REGION Network 75
   RUNG wire#powerrail
      Contact( "LimiteMantBoost2" )
      Coil( "DB32".Static_194 )
   END_RUNG
   // the same network as SCL:
   "DB32".Static_194 := "LimiteMantBoost2";
END_REGION

REGION Network 76
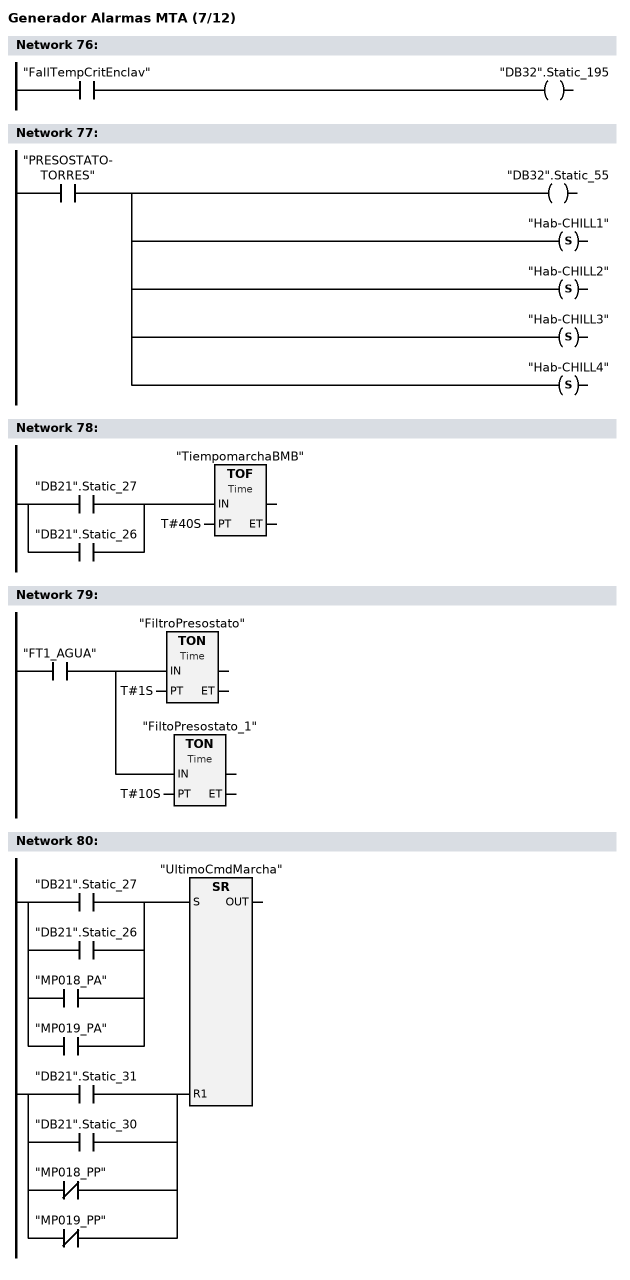
   RUNG wire#powerrail
      Contact( "FallTempCritEnclav" )
      Coil( "DB32".Static_195 )
   END_RUNG
   // the same network as SCL:
   "DB32".Static_195 := "FallTempCritEnclav";
END_REGION

REGION Network 77
   RUNG wire#powerrail
      Contact( "PRESOSTATO-TORRES" )
      wire#w1
      Coil( "DB32".Static_55 )
   END_RUNG
   RUNG wire#w1
      S_Coil( "Hab-CHILL1" )
   END_RUNG
   RUNG wire#w1
      S_Coil( "Hab-CHILL2" )
   END_RUNG
   RUNG wire#w1
      S_Coil( "Hab-CHILL3" )
   END_RUNG
   RUNG wire#w1
      S_Coil( "Hab-CHILL4" )
   END_RUNG
   // the same network as SCL:
   "DB32".Static_55 := "PRESOSTATO-TORRES";
   IF "PRESOSTATO-TORRES" THEN
       "Hab-CHILL1" := TRUE;
       "Hab-CHILL2" := TRUE;
       "Hab-CHILL3" := TRUE;
       "Hab-CHILL4" := TRUE;
   END_IF;
END_REGION

REGION Network 78
   "TiempomarchaBMB".TOF(in := "DB21".Static_27 OR "DB21".Static_26, pt := T#40S);
END_REGION

REGION Network 79
   "FiltroPresostato".TON(pt := T#1S, in := "FT1_AGUA");
   "FiltoPresostato_1".TON(pt := T#10S, in := "FT1_AGUA");
END_REGION

REGION Network 80
   RUNG wire#powerrail
      Contact( "DB21".Static_27 )
      wire#w1
      S_SR(operand := "UltimoCmdMarcha", r1 := wire#w2)
   END_RUNG
   RUNG wire#powerrail
      Contact( "DB21".Static_26 )
   END_RUNG wire#w1
   RUNG wire#powerrail
      Contact( "MP018_PA" )
   END_RUNG wire#w1
   RUNG wire#powerrail
      Contact( "MP019_PA" )
   END_RUNG wire#w1
   RUNG wire#powerrail
      Contact( "DB21".Static_31 )
   END_RUNG wire#w2
   RUNG wire#powerrail
      Contact( "DB21".Static_30 )
   END_RUNG wire#w2
   RUNG wire#powerrail
      I_Contact( "MP018_PP" )
   END_RUNG wire#w2
   RUNG wire#powerrail
      I_Contact( "MP019_PP" )
   END_RUNG wire#w2
   // the same network as SCL:
   IF "DB21".Static_27 OR "DB21".Static_26 OR "MP018_PA" OR "MP019_PA" THEN
       "UltimoCmdMarcha" := TRUE;   // SR flip-flop
   END_IF;
   IF "DB21".Static_31 OR "DB21".Static_30 OR NOT "MP018_PP" OR NOT "MP019_PP" THEN
       "UltimoCmdMarcha" := FALSE;
   END_IF;
END_REGION

REGION Network 81
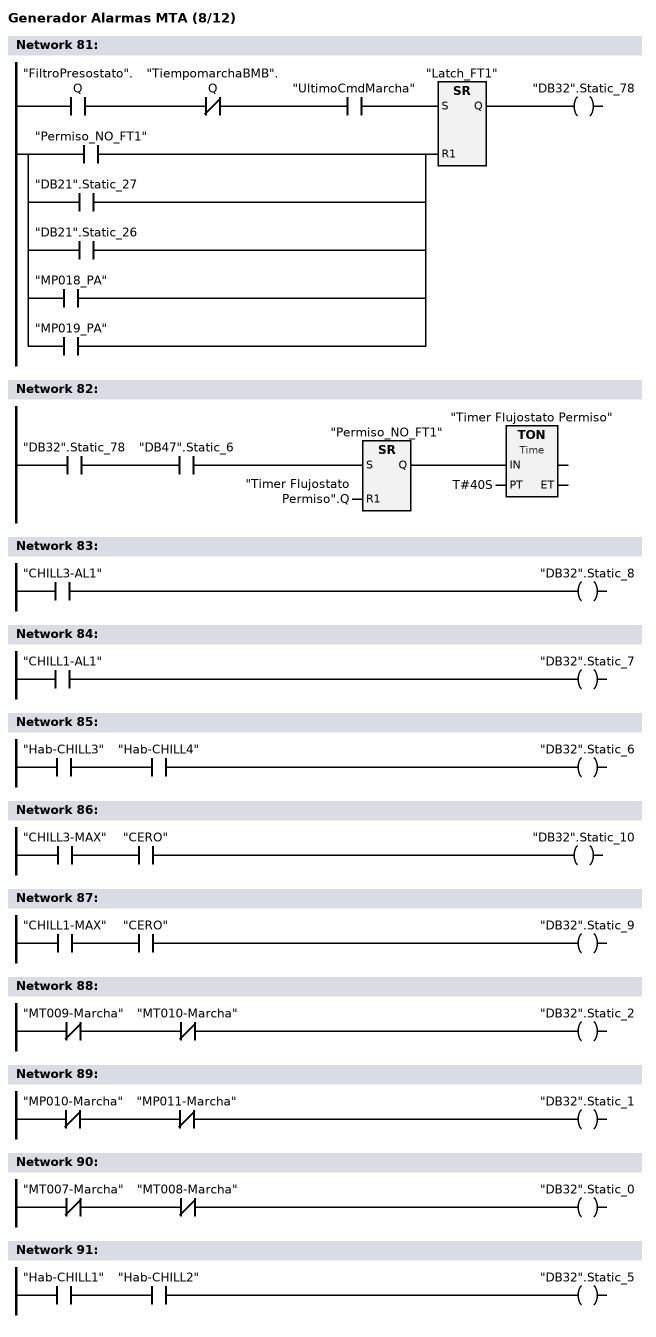
   RUNG wire#powerrail
      Contact( "FiltroPresostato".Q )
      I_Contact( "TiempomarchaBMB".Q )
      Contact( "UltimoCmdMarcha" )
      S_SR(operand := "Latch_FT1", r1 := wire#w1)
      Coil( "DB32".Static_78 )
   END_RUNG
   RUNG wire#powerrail
      Contact( "Permiso_NO_FT1" )
   END_RUNG wire#w1
   RUNG wire#powerrail
      Contact( "DB21".Static_27 )
   END_RUNG wire#w1
   RUNG wire#powerrail
      Contact( "DB21".Static_26 )
   END_RUNG wire#w1
   RUNG wire#powerrail
      Contact( "MP018_PA" )
   END_RUNG wire#w1
   RUNG wire#powerrail
      Contact( "MP019_PA" )
   END_RUNG wire#w1
   // the same network as SCL:
   IF "FiltroPresostato".Q AND NOT "TiempomarchaBMB".Q AND "UltimoCmdMarcha" THEN
       "Latch_FT1" := TRUE;   // SR flip-flop
   END_IF;
   IF "Permiso_NO_FT1" OR "DB21".Static_27 OR "DB21".Static_26 OR "MP018_PA" OR "MP019_PA" THEN
       "Latch_FT1" := FALSE;
   END_IF;
   "DB32".Static_78 := "Latch_FT1";
END_REGION

REGION Network 82
   IF "DB32".Static_78 AND "DB47".Static_6 THEN
       "Permiso_NO_FT1" := TRUE;   // SR flip-flop
   END_IF;
   IF "Timer Flujostato Permiso".Q THEN "Permiso_NO_FT1" := FALSE; END_IF;
   "Timer Flujostato Permiso".TON(in := "Permiso_NO_FT1", pt := T#40S);
END_REGION

REGION Network 83
   RUNG wire#powerrail
      Contact( "CHILL3-AL1" )
      Coil( "DB32".Static_8 )
   END_RUNG
   // the same network as SCL:
   "DB32".Static_8 := "CHILL3-AL1";
END_REGION

REGION Network 84
   RUNG wire#powerrail
      Contact( "CHILL1-AL1" )
      Coil( "DB32".Static_7 )
   END_RUNG
   // the same network as SCL:
   "DB32".Static_7 := "CHILL1-AL1";
END_REGION

REGION Network 85
   RUNG wire#powerrail
      Contact( "Hab-CHILL3" )
      Contact( "Hab-CHILL4" )
      Coil( "DB32".Static_6 )
   END_RUNG
   // the same network as SCL:
   "DB32".Static_6 := "Hab-CHILL3" AND "Hab-CHILL4";
END_REGION

REGION Network 86
   RUNG wire#powerrail
      Contact( "CHILL3-MAX" )
      Contact( "CERO" )
      Coil( "DB32".Static_10 )
   END_RUNG
   // the same network as SCL:
   "DB32".Static_10 := "CHILL3-MAX" AND "CERO";
END_REGION

REGION Network 87
   RUNG wire#powerrail
      Contact( "CHILL1-MAX" )
      Contact( "CERO" )
      Coil( "DB32".Static_9 )
   END_RUNG
   // the same network as SCL:
   "DB32".Static_9 := "CHILL1-MAX" AND "CERO";
END_REGION

REGION Network 88
   RUNG wire#powerrail
      I_Contact( "MT009-Marcha" )
      I_Contact( "MT010-Marcha" )
      Coil( "DB32".Static_2 )
   END_RUNG
   // the same network as SCL:
   "DB32".Static_2 := NOT "MT009-Marcha" AND NOT "MT010-Marcha";
END_REGION

REGION Network 89
   RUNG wire#powerrail
      I_Contact( "MP010-Marcha" )
      I_Contact( "MP011-Marcha" )
      Coil( "DB32".Static_1 )
   END_RUNG
   // the same network as SCL:
   "DB32".Static_1 := NOT "MP010-Marcha" AND NOT "MP011-Marcha";
END_REGION

REGION Network 90
   RUNG wire#powerrail
      I_Contact( "MT007-Marcha" )
      I_Contact( "MT008-Marcha" )
      Coil( "DB32".Static_0 )
   END_RUNG
   // the same network as SCL:
   "DB32".Static_0 := NOT "MT007-Marcha" AND NOT "MT008-Marcha";
END_REGION

REGION Network 91
   RUNG wire#powerrail
      Contact( "Hab-CHILL1" )
      Contact( "Hab-CHILL2" )
      Coil( "DB32".Static_5 )
   END_RUNG
   // the same network as SCL:
   "DB32".Static_5 := "Hab-CHILL1" AND "Hab-CHILL2";
END_REGION

REGION Network 92
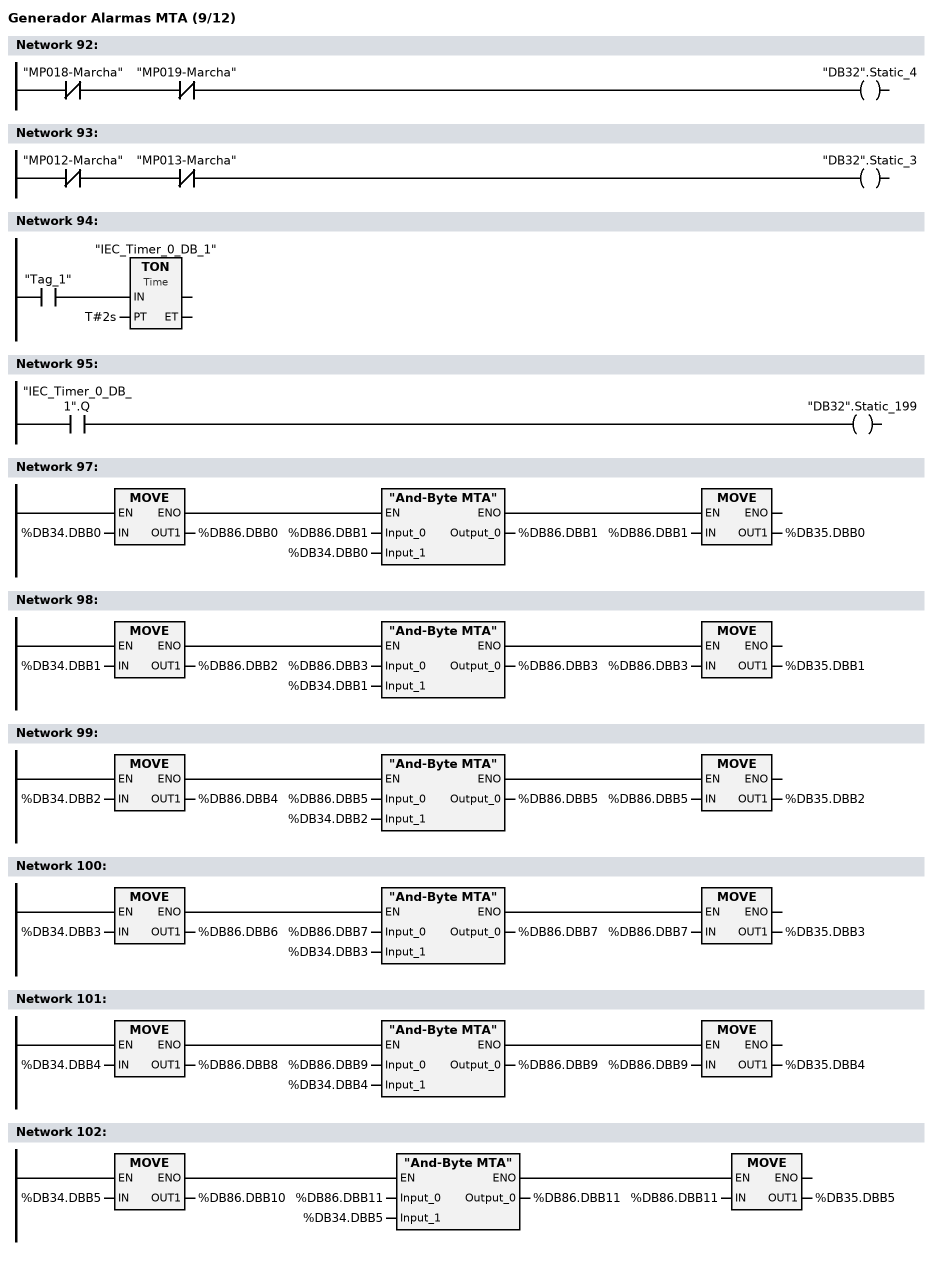
   RUNG wire#powerrail
      I_Contact( "MP018-Marcha" )
      I_Contact( "MP019-Marcha" )
      Coil( "DB32".Static_4 )
   END_RUNG
   // the same network as SCL:
   "DB32".Static_4 := NOT "MP018-Marcha" AND NOT "MP019-Marcha";
END_REGION

REGION Network 93
   RUNG wire#powerrail
      I_Contact( "MP012-Marcha" )
      I_Contact( "MP013-Marcha" )
      Coil( "DB32".Static_3 )
   END_RUNG
   // the same network as SCL:
   "DB32".Static_3 := NOT "MP012-Marcha" AND NOT "MP013-Marcha";
END_REGION

REGION Network 94
   "IEC_Timer_0_DB_1".TON(IN := "Tag_1", PT := T#2s);
END_REGION

REGION Network 95
   RUNG wire#powerrail
      Contact( "IEC_Timer_0_DB_1".Q )
      Coil( "DB32".Static_199 )
   END_RUNG
   // the same network as SCL:
   "DB32".Static_199 := "IEC_Timer_0_DB_1".Q;
END_REGION

REGION Network 97
   RUNG wire#powerrail
      { S7_GenerateENO := "TRUE" } Move(in := %DB34.DBB0, out1 => %DB86.DBB0)
      "And-Byte MTA"(Input_0 := %DB86.DBB1, Input_1 := %DB34.DBB0, Output_0 => %DB86.DBB1)
      { S7_GenerateENO := "TRUE" } Move(in := %DB86.DBB1, out1 => %DB35.DBB0)
   END_RUNG
   // the same network as SCL:
   // ENO of a box is taken as its EN; it also drops when the box reports an error
   %DB86.DBB0 := %DB34.DBB0;
   "And-Byte MTA"(Input_0 := %DB86.DBB1, Input_1 := %DB34.DBB0, Output_0 => %DB86.DBB1, ENO => #_w1);
   IF #_w1 THEN %DB35.DBB0 := %DB86.DBB1; END_IF;
END_REGION

REGION Network 98
   RUNG wire#powerrail
      { S7_GenerateENO := "TRUE" } Move(in := %DB34.DBB1, out1 => %DB86.DBB2)
      "And-Byte MTA"(Input_0 := %DB86.DBB3, Input_1 := %DB34.DBB1, Output_0 => %DB86.DBB3)
      { S7_GenerateENO := "TRUE" } Move(in := %DB86.DBB3, out1 => %DB35.DBB1)
   END_RUNG
   // the same network as SCL:
   // ENO of a box is taken as its EN; it also drops when the box reports an error
   %DB86.DBB2 := %DB34.DBB1;
   "And-Byte MTA"(Input_0 := %DB86.DBB3, Input_1 := %DB34.DBB1, Output_0 => %DB86.DBB3, ENO => #_w1);
   IF #_w1 THEN %DB35.DBB1 := %DB86.DBB3; END_IF;
END_REGION

REGION Network 99
   RUNG wire#powerrail
      { S7_GenerateENO := "TRUE" } Move(in := %DB34.DBB2, out1 => %DB86.DBB4)
      "And-Byte MTA"(Input_0 := %DB86.DBB5, Input_1 := %DB34.DBB2, Output_0 => %DB86.DBB5)
      { S7_GenerateENO := "TRUE" } Move(in := %DB86.DBB5, out1 => %DB35.DBB2)
   END_RUNG
   // the same network as SCL:
   // ENO of a box is taken as its EN; it also drops when the box reports an error
   %DB86.DBB4 := %DB34.DBB2;
   "And-Byte MTA"(Input_0 := %DB86.DBB5, Input_1 := %DB34.DBB2, Output_0 => %DB86.DBB5, ENO => #_w1);
   IF #_w1 THEN %DB35.DBB2 := %DB86.DBB5; END_IF;
END_REGION

REGION Network 100
   RUNG wire#powerrail
      { S7_GenerateENO := "TRUE" } Move(in := %DB34.DBB3, out1 => %DB86.DBB6)
      "And-Byte MTA"(Input_0 := %DB86.DBB7, Input_1 := %DB34.DBB3, Output_0 => %DB86.DBB7)
      { S7_GenerateENO := "TRUE" } Move(in := %DB86.DBB7, out1 => %DB35.DBB3)
   END_RUNG
   // the same network as SCL:
   // ENO of a box is taken as its EN; it also drops when the box reports an error
   %DB86.DBB6 := %DB34.DBB3;
   "And-Byte MTA"(Input_0 := %DB86.DBB7, Input_1 := %DB34.DBB3, Output_0 => %DB86.DBB7, ENO => #_w1);
   IF #_w1 THEN %DB35.DBB3 := %DB86.DBB7; END_IF;
END_REGION

REGION Network 101
   RUNG wire#powerrail
      { S7_GenerateENO := "TRUE" } Move(in := %DB34.DBB4, out1 => %DB86.DBB8)
      "And-Byte MTA"(Input_0 := %DB86.DBB9, Input_1 := %DB34.DBB4, Output_0 => %DB86.DBB9)
      { S7_GenerateENO := "TRUE" } Move(in := %DB86.DBB9, out1 => %DB35.DBB4)
   END_RUNG
   // the same network as SCL:
   // ENO of a box is taken as its EN; it also drops when the box reports an error
   %DB86.DBB8 := %DB34.DBB4;
   "And-Byte MTA"(Input_0 := %DB86.DBB9, Input_1 := %DB34.DBB4, Output_0 => %DB86.DBB9, ENO => #_w1);
   IF #_w1 THEN %DB35.DBB4 := %DB86.DBB9; END_IF;
END_REGION

REGION Network 102
   RUNG wire#powerrail
      { S7_GenerateENO := "TRUE" } Move(in := %DB34.DBB5, out1 => %DB86.DBB10)
      "And-Byte MTA"(Input_0 := %DB86.DBB11, Input_1 := %DB34.DBB5, Output_0 => %DB86.DBB11)
      { S7_GenerateENO := "TRUE" } Move(in := %DB86.DBB11, out1 => %DB35.DBB5)
   END_RUNG
   // the same network as SCL:
   // ENO of a box is taken as its EN; it also drops when the box reports an error
   %DB86.DBB10 := %DB34.DBB5;
   "And-Byte MTA"(Input_0 := %DB86.DBB11, Input_1 := %DB34.DBB5, Output_0 => %DB86.DBB11, ENO => #_w1);
   IF #_w1 THEN %DB35.DBB5 := %DB86.DBB11; END_IF;
END_REGION

REGION Network 103
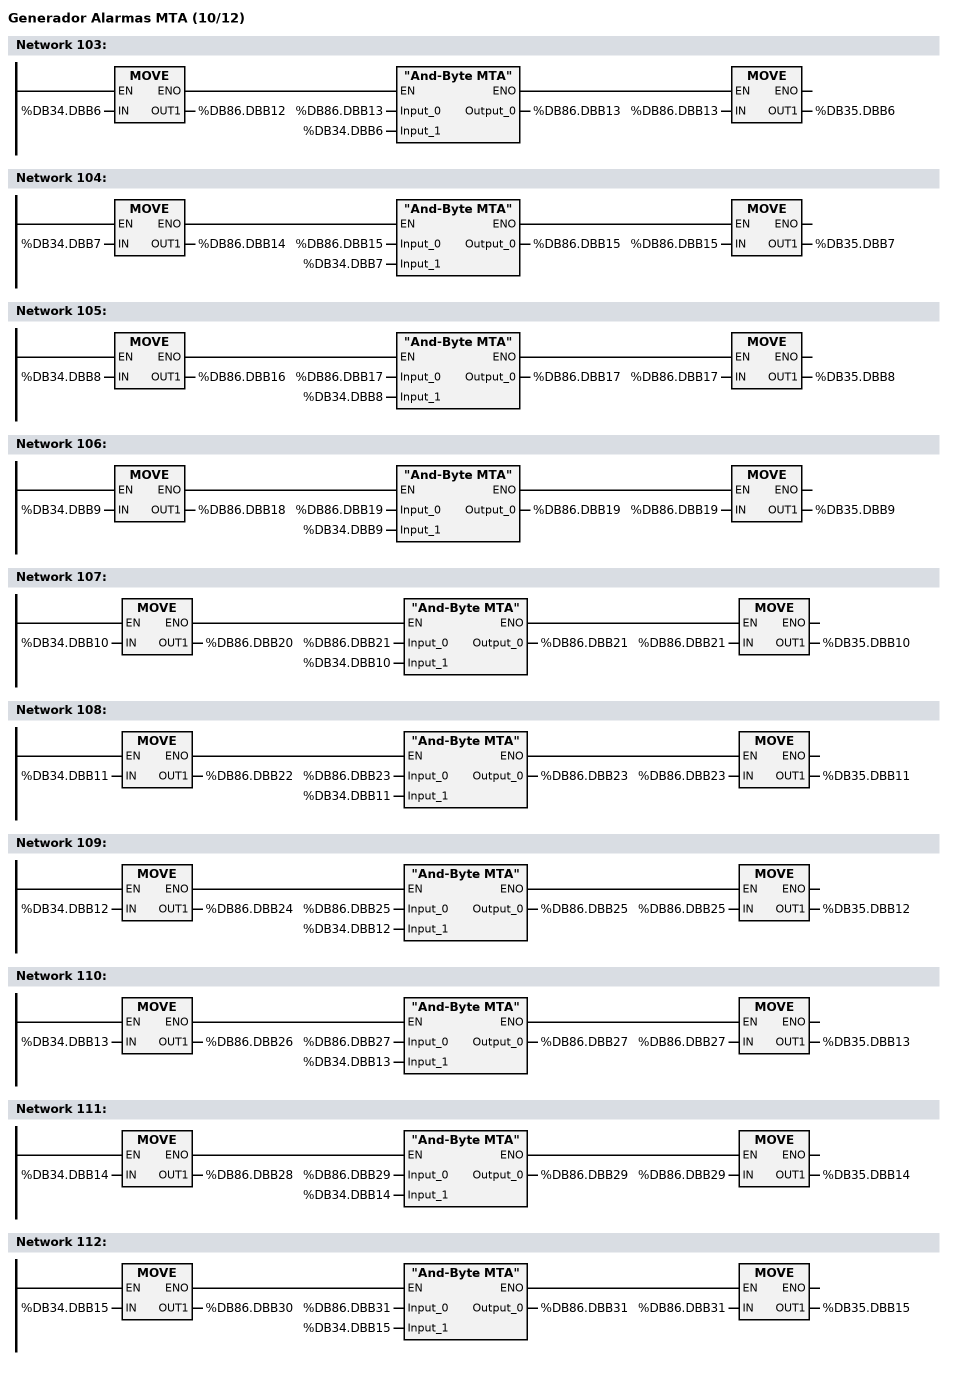
   RUNG wire#powerrail
      { S7_GenerateENO := "TRUE" } Move(in := %DB34.DBB6, out1 => %DB86.DBB12)
      "And-Byte MTA"(Input_0 := %DB86.DBB13, Input_1 := %DB34.DBB6, Output_0 => %DB86.DBB13)
      { S7_GenerateENO := "TRUE" } Move(in := %DB86.DBB13, out1 => %DB35.DBB6)
   END_RUNG
   // the same network as SCL:
   // ENO of a box is taken as its EN; it also drops when the box reports an error
   %DB86.DBB12 := %DB34.DBB6;
   "And-Byte MTA"(Input_0 := %DB86.DBB13, Input_1 := %DB34.DBB6, Output_0 => %DB86.DBB13, ENO => #_w1);
   IF #_w1 THEN %DB35.DBB6 := %DB86.DBB13; END_IF;
END_REGION

REGION Network 104
   RUNG wire#powerrail
      { S7_GenerateENO := "TRUE" } Move(in := %DB34.DBB7, out1 => %DB86.DBB14)
      "And-Byte MTA"(Input_0 := %DB86.DBB15, Input_1 := %DB34.DBB7, Output_0 => %DB86.DBB15)
      { S7_GenerateENO := "TRUE" } Move(in := %DB86.DBB15, out1 => %DB35.DBB7)
   END_RUNG
   // the same network as SCL:
   // ENO of a box is taken as its EN; it also drops when the box reports an error
   %DB86.DBB14 := %DB34.DBB7;
   "And-Byte MTA"(Input_0 := %DB86.DBB15, Input_1 := %DB34.DBB7, Output_0 => %DB86.DBB15, ENO => #_w1);
   IF #_w1 THEN %DB35.DBB7 := %DB86.DBB15; END_IF;
END_REGION

REGION Network 105
   RUNG wire#powerrail
      { S7_GenerateENO := "TRUE" } Move(in := %DB34.DBB8, out1 => %DB86.DBB16)
      "And-Byte MTA"(Input_0 := %DB86.DBB17, Input_1 := %DB34.DBB8, Output_0 => %DB86.DBB17)
      { S7_GenerateENO := "TRUE" } Move(in := %DB86.DBB17, out1 => %DB35.DBB8)
   END_RUNG
   // the same network as SCL:
   // ENO of a box is taken as its EN; it also drops when the box reports an error
   %DB86.DBB16 := %DB34.DBB8;
   "And-Byte MTA"(Input_0 := %DB86.DBB17, Input_1 := %DB34.DBB8, Output_0 => %DB86.DBB17, ENO => #_w1);
   IF #_w1 THEN %DB35.DBB8 := %DB86.DBB17; END_IF;
END_REGION

REGION Network 106
   RUNG wire#powerrail
      { S7_GenerateENO := "TRUE" } Move(in := %DB34.DBB9, out1 => %DB86.DBB18)
      "And-Byte MTA"(Input_0 := %DB86.DBB19, Input_1 := %DB34.DBB9, Output_0 => %DB86.DBB19)
      { S7_GenerateENO := "TRUE" } Move(in := %DB86.DBB19, out1 => %DB35.DBB9)
   END_RUNG
   // the same network as SCL:
   // ENO of a box is taken as its EN; it also drops when the box reports an error
   %DB86.DBB18 := %DB34.DBB9;
   "And-Byte MTA"(Input_0 := %DB86.DBB19, Input_1 := %DB34.DBB9, Output_0 => %DB86.DBB19, ENO => #_w1);
   IF #_w1 THEN %DB35.DBB9 := %DB86.DBB19; END_IF;
END_REGION

REGION Network 107
   RUNG wire#powerrail
      { S7_GenerateENO := "TRUE" } Move(in := %DB34.DBB10, out1 => %DB86.DBB20)
      "And-Byte MTA"(Input_0 := %DB86.DBB21, Input_1 := %DB34.DBB10, Output_0 => %DB86.DBB21)
      { S7_GenerateENO := "TRUE" } Move(in := %DB86.DBB21, out1 => %DB35.DBB10)
   END_RUNG
   // the same network as SCL:
   // ENO of a box is taken as its EN; it also drops when the box reports an error
   %DB86.DBB20 := %DB34.DBB10;
   "And-Byte MTA"(Input_0 := %DB86.DBB21, Input_1 := %DB34.DBB10, Output_0 => %DB86.DBB21, ENO => #_w1);
   IF #_w1 THEN %DB35.DBB10 := %DB86.DBB21; END_IF;
END_REGION

REGION Network 108
   RUNG wire#powerrail
      { S7_GenerateENO := "TRUE" } Move(in := %DB34.DBB11, out1 => %DB86.DBB22)
      "And-Byte MTA"(Input_0 := %DB86.DBB23, Input_1 := %DB34.DBB11, Output_0 => %DB86.DBB23)
      { S7_GenerateENO := "TRUE" } Move(in := %DB86.DBB23, out1 => %DB35.DBB11)
   END_RUNG
   // the same network as SCL:
   // ENO of a box is taken as its EN; it also drops when the box reports an error
   %DB86.DBB22 := %DB34.DBB11;
   "And-Byte MTA"(Input_0 := %DB86.DBB23, Input_1 := %DB34.DBB11, Output_0 => %DB86.DBB23, ENO => #_w1);
   IF #_w1 THEN %DB35.DBB11 := %DB86.DBB23; END_IF;
END_REGION

REGION Network 109
   RUNG wire#powerrail
      { S7_GenerateENO := "TRUE" } Move(in := %DB34.DBB12, out1 => %DB86.DBB24)
      "And-Byte MTA"(Input_0 := %DB86.DBB25, Input_1 := %DB34.DBB12, Output_0 => %DB86.DBB25)
      { S7_GenerateENO := "TRUE" } Move(in := %DB86.DBB25, out1 => %DB35.DBB12)
   END_RUNG
   // the same network as SCL:
   // ENO of a box is taken as its EN; it also drops when the box reports an error
   %DB86.DBB24 := %DB34.DBB12;
   "And-Byte MTA"(Input_0 := %DB86.DBB25, Input_1 := %DB34.DBB12, Output_0 => %DB86.DBB25, ENO => #_w1);
   IF #_w1 THEN %DB35.DBB12 := %DB86.DBB25; END_IF;
END_REGION

REGION Network 110
   RUNG wire#powerrail
      { S7_GenerateENO := "TRUE" } Move(in := %DB34.DBB13, out1 => %DB86.DBB26)
      "And-Byte MTA"(Input_0 := %DB86.DBB27, Input_1 := %DB34.DBB13, Output_0 => %DB86.DBB27)
      { S7_GenerateENO := "TRUE" } Move(in := %DB86.DBB27, out1 => %DB35.DBB13)
   END_RUNG
   // the same network as SCL:
   // ENO of a box is taken as its EN; it also drops when the box reports an error
   %DB86.DBB26 := %DB34.DBB13;
   "And-Byte MTA"(Input_0 := %DB86.DBB27, Input_1 := %DB34.DBB13, Output_0 => %DB86.DBB27, ENO => #_w1);
   IF #_w1 THEN %DB35.DBB13 := %DB86.DBB27; END_IF;
END_REGION

REGION Network 111
   RUNG wire#powerrail
      { S7_GenerateENO := "TRUE" } Move(in := %DB34.DBB14, out1 => %DB86.DBB28)
      "And-Byte MTA"(Input_0 := %DB86.DBB29, Input_1 := %DB34.DBB14, Output_0 => %DB86.DBB29)
      { S7_GenerateENO := "TRUE" } Move(in := %DB86.DBB29, out1 => %DB35.DBB14)
   END_RUNG
   // the same network as SCL:
   // ENO of a box is taken as its EN; it also drops when the box reports an error
   %DB86.DBB28 := %DB34.DBB14;
   "And-Byte MTA"(Input_0 := %DB86.DBB29, Input_1 := %DB34.DBB14, Output_0 => %DB86.DBB29, ENO => #_w1);
   IF #_w1 THEN %DB35.DBB14 := %DB86.DBB29; END_IF;
END_REGION

REGION Network 112
   RUNG wire#powerrail
      { S7_GenerateENO := "TRUE" } Move(in := %DB34.DBB15, out1 => %DB86.DBB30)
      "And-Byte MTA"(Input_0 := %DB86.DBB31, Input_1 := %DB34.DBB15, Output_0 => %DB86.DBB31)
      { S7_GenerateENO := "TRUE" } Move(in := %DB86.DBB31, out1 => %DB35.DBB15)
   END_RUNG
   // the same network as SCL:
   // ENO of a box is taken as its EN; it also drops when the box reports an error
   %DB86.DBB30 := %DB34.DBB15;
   "And-Byte MTA"(Input_0 := %DB86.DBB31, Input_1 := %DB34.DBB15, Output_0 => %DB86.DBB31, ENO => #_w1);
   IF #_w1 THEN %DB35.DBB15 := %DB86.DBB31; END_IF;
END_REGION

REGION Network 113
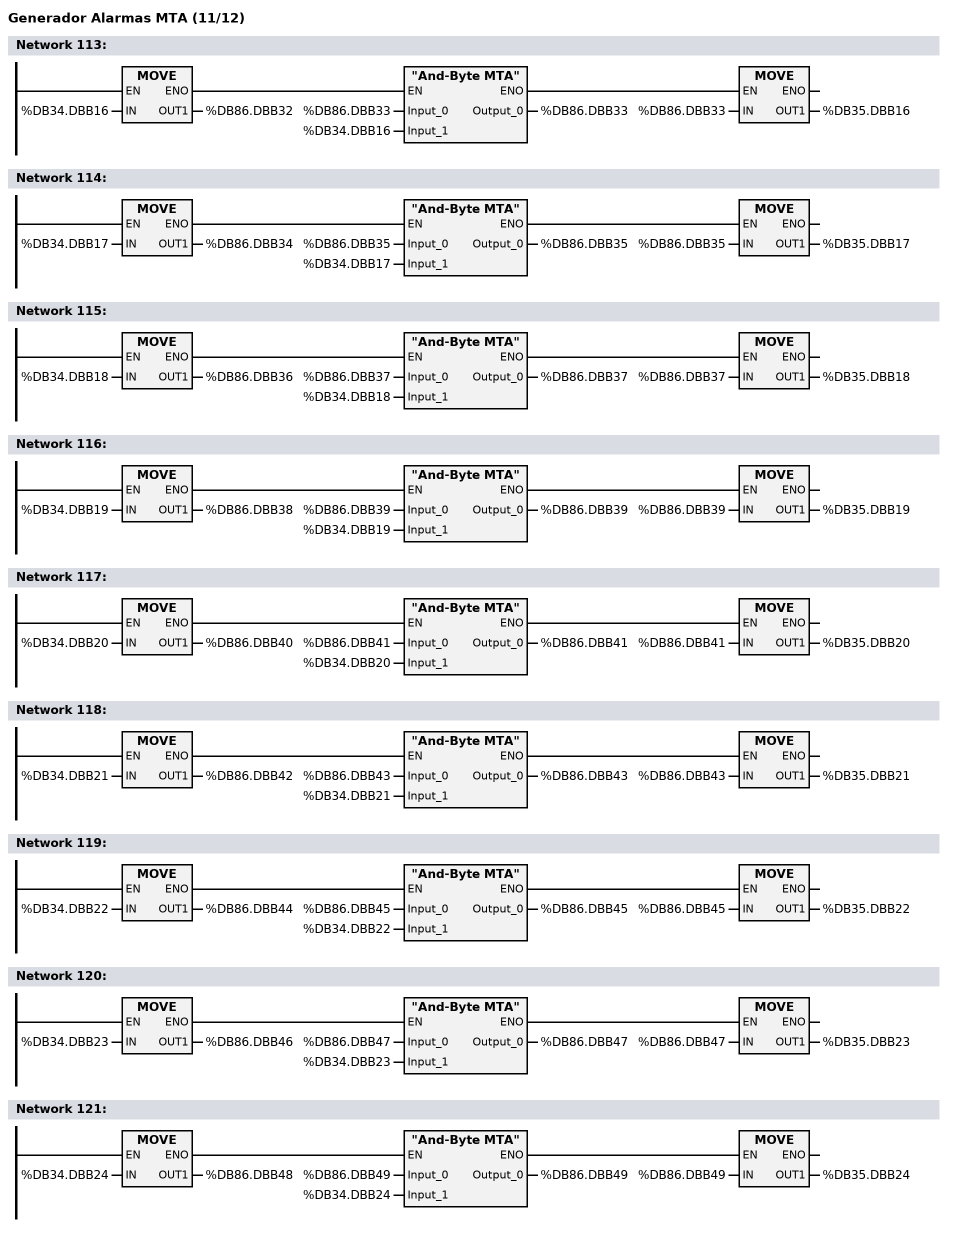
   RUNG wire#powerrail
      { S7_GenerateENO := "TRUE" } Move(in := %DB34.DBB16, out1 => %DB86.DBB32)
      "And-Byte MTA"(Input_0 := %DB86.DBB33, Input_1 := %DB34.DBB16, Output_0 => %DB86.DBB33)
      { S7_GenerateENO := "TRUE" } Move(in := %DB86.DBB33, out1 => %DB35.DBB16)
   END_RUNG
   // the same network as SCL:
   // ENO of a box is taken as its EN; it also drops when the box reports an error
   %DB86.DBB32 := %DB34.DBB16;
   "And-Byte MTA"(Input_0 := %DB86.DBB33, Input_1 := %DB34.DBB16, Output_0 => %DB86.DBB33, ENO => #_w1);
   IF #_w1 THEN %DB35.DBB16 := %DB86.DBB33; END_IF;
END_REGION

REGION Network 114
   RUNG wire#powerrail
      { S7_GenerateENO := "TRUE" } Move(in := %DB34.DBB17, out1 => %DB86.DBB34)
      "And-Byte MTA"(Input_0 := %DB86.DBB35, Input_1 := %DB34.DBB17, Output_0 => %DB86.DBB35)
      { S7_GenerateENO := "TRUE" } Move(in := %DB86.DBB35, out1 => %DB35.DBB17)
   END_RUNG
   // the same network as SCL:
   // ENO of a box is taken as its EN; it also drops when the box reports an error
   %DB86.DBB34 := %DB34.DBB17;
   "And-Byte MTA"(Input_0 := %DB86.DBB35, Input_1 := %DB34.DBB17, Output_0 => %DB86.DBB35, ENO => #_w1);
   IF #_w1 THEN %DB35.DBB17 := %DB86.DBB35; END_IF;
END_REGION

REGION Network 115
   RUNG wire#powerrail
      { S7_GenerateENO := "TRUE" } Move(in := %DB34.DBB18, out1 => %DB86.DBB36)
      "And-Byte MTA"(Input_0 := %DB86.DBB37, Input_1 := %DB34.DBB18, Output_0 => %DB86.DBB37)
      { S7_GenerateENO := "TRUE" } Move(in := %DB86.DBB37, out1 => %DB35.DBB18)
   END_RUNG
   // the same network as SCL:
   // ENO of a box is taken as its EN; it also drops when the box reports an error
   %DB86.DBB36 := %DB34.DBB18;
   "And-Byte MTA"(Input_0 := %DB86.DBB37, Input_1 := %DB34.DBB18, Output_0 => %DB86.DBB37, ENO => #_w1);
   IF #_w1 THEN %DB35.DBB18 := %DB86.DBB37; END_IF;
END_REGION

REGION Network 116
   RUNG wire#powerrail
      { S7_GenerateENO := "TRUE" } Move(in := %DB34.DBB19, out1 => %DB86.DBB38)
      "And-Byte MTA"(Input_0 := %DB86.DBB39, Input_1 := %DB34.DBB19, Output_0 => %DB86.DBB39)
      { S7_GenerateENO := "TRUE" } Move(in := %DB86.DBB39, out1 => %DB35.DBB19)
   END_RUNG
   // the same network as SCL:
   // ENO of a box is taken as its EN; it also drops when the box reports an error
   %DB86.DBB38 := %DB34.DBB19;
   "And-Byte MTA"(Input_0 := %DB86.DBB39, Input_1 := %DB34.DBB19, Output_0 => %DB86.DBB39, ENO => #_w1);
   IF #_w1 THEN %DB35.DBB19 := %DB86.DBB39; END_IF;
END_REGION

REGION Network 117
   RUNG wire#powerrail
      { S7_GenerateENO := "TRUE" } Move(in := %DB34.DBB20, out1 => %DB86.DBB40)
      "And-Byte MTA"(Input_0 := %DB86.DBB41, Input_1 := %DB34.DBB20, Output_0 => %DB86.DBB41)
      { S7_GenerateENO := "TRUE" } Move(in := %DB86.DBB41, out1 => %DB35.DBB20)
   END_RUNG
   // the same network as SCL:
   // ENO of a box is taken as its EN; it also drops when the box reports an error
   %DB86.DBB40 := %DB34.DBB20;
   "And-Byte MTA"(Input_0 := %DB86.DBB41, Input_1 := %DB34.DBB20, Output_0 => %DB86.DBB41, ENO => #_w1);
   IF #_w1 THEN %DB35.DBB20 := %DB86.DBB41; END_IF;
END_REGION

REGION Network 118
   RUNG wire#powerrail
      { S7_GenerateENO := "TRUE" } Move(in := %DB34.DBB21, out1 => %DB86.DBB42)
      "And-Byte MTA"(Input_0 := %DB86.DBB43, Input_1 := %DB34.DBB21, Output_0 => %DB86.DBB43)
      { S7_GenerateENO := "TRUE" } Move(in := %DB86.DBB43, out1 => %DB35.DBB21)
   END_RUNG
   // the same network as SCL:
   // ENO of a box is taken as its EN; it also drops when the box reports an error
   %DB86.DBB42 := %DB34.DBB21;
   "And-Byte MTA"(Input_0 := %DB86.DBB43, Input_1 := %DB34.DBB21, Output_0 => %DB86.DBB43, ENO => #_w1);
   IF #_w1 THEN %DB35.DBB21 := %DB86.DBB43; END_IF;
END_REGION

REGION Network 119
   RUNG wire#powerrail
      { S7_GenerateENO := "TRUE" } Move(in := %DB34.DBB22, out1 => %DB86.DBB44)
      "And-Byte MTA"(Input_0 := %DB86.DBB45, Input_1 := %DB34.DBB22, Output_0 => %DB86.DBB45)
      { S7_GenerateENO := "TRUE" } Move(in := %DB86.DBB45, out1 => %DB35.DBB22)
   END_RUNG
   // the same network as SCL:
   // ENO of a box is taken as its EN; it also drops when the box reports an error
   %DB86.DBB44 := %DB34.DBB22;
   "And-Byte MTA"(Input_0 := %DB86.DBB45, Input_1 := %DB34.DBB22, Output_0 => %DB86.DBB45, ENO => #_w1);
   IF #_w1 THEN %DB35.DBB22 := %DB86.DBB45; END_IF;
END_REGION

REGION Network 120
   RUNG wire#powerrail
      { S7_GenerateENO := "TRUE" } Move(in := %DB34.DBB23, out1 => %DB86.DBB46)
      "And-Byte MTA"(Input_0 := %DB86.DBB47, Input_1 := %DB34.DBB23, Output_0 => %DB86.DBB47)
      { S7_GenerateENO := "TRUE" } Move(in := %DB86.DBB47, out1 => %DB35.DBB23)
   END_RUNG
   // the same network as SCL:
   // ENO of a box is taken as its EN; it also drops when the box reports an error
   %DB86.DBB46 := %DB34.DBB23;
   "And-Byte MTA"(Input_0 := %DB86.DBB47, Input_1 := %DB34.DBB23, Output_0 => %DB86.DBB47, ENO => #_w1);
   IF #_w1 THEN %DB35.DBB23 := %DB86.DBB47; END_IF;
END_REGION

REGION Network 121
   RUNG wire#powerrail
      { S7_GenerateENO := "TRUE" } Move(in := %DB34.DBB24, out1 => %DB86.DBB48)
      "And-Byte MTA"(Input_0 := %DB86.DBB49, Input_1 := %DB34.DBB24, Output_0 => %DB86.DBB49)
      { S7_GenerateENO := "TRUE" } Move(in := %DB86.DBB49, out1 => %DB35.DBB24)
   END_RUNG
   // the same network as SCL:
   // ENO of a box is taken as its EN; it also drops when the box reports an error
   %DB86.DBB48 := %DB34.DBB24;
   "And-Byte MTA"(Input_0 := %DB86.DBB49, Input_1 := %DB34.DBB24, Output_0 => %DB86.DBB49, ENO => #_w1);
   IF #_w1 THEN %DB35.DBB24 := %DB86.DBB49; END_IF;
END_REGION

REGION Network 122
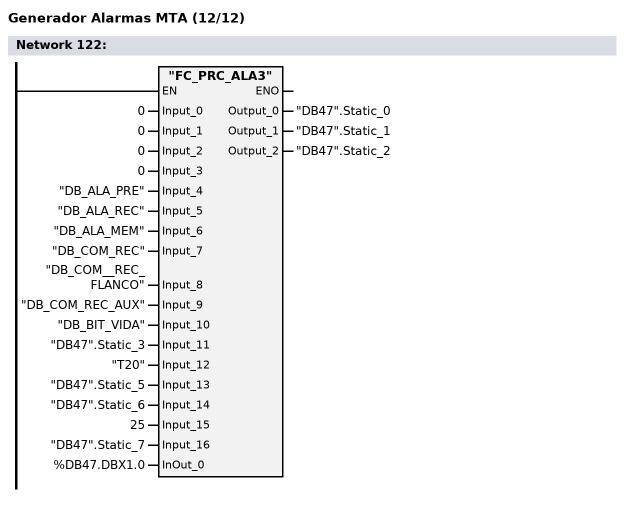
   RUNG wire#powerrail
      "FC_PRC_ALA3"(Input_0 := 0, Input_1 := 0, Input_2 := 0, Input_3 := 0, Input_4 := "DB_ALA_PRE", Input_5 := "DB_ALA_REC", Input_6 := "DB_ALA_MEM", Input_7 := "DB_COM_REC", Input_8 := "DB_COM__REC_FLANCO", Input_9 := "DB_COM_REC_AUX", Input_10 := "DB_BIT_VIDA", Input_11 := "DB47".Static_3, Input_12 := "T20", Input_13 := "DB47".Static_5, Input_14 := "DB47".Static_6, Input_15 := 25, Input_16 := "DB47".Static_7, Output_0 => "DB47".Static_0, Output_1 => "DB47".Static_1, Output_2 => "DB47".Static_2, InOut_0 := %DB47.DBX1.0)
   END_RUNG
   // the same network as SCL:
   "FC_PRC_ALA3"(Input_0 := 0,
                 Input_1 := 0,
                 Input_2 := 0,
                 Input_3 := 0,
                 Input_4 := "DB_ALA_PRE",
                 Input_5 := "DB_ALA_REC",
                 Input_6 := "DB_ALA_MEM",
                 Input_7 := "DB_COM_REC",
                 Input_8 := "DB_COM__REC_FLANCO",
                 Input_9 := "DB_COM_REC_AUX",
                 Input_10 := "DB_BIT_VIDA",
                 Input_11 := "DB47".Static_3,
                 Input_12 := "T20",
                 Input_13 := "DB47".Static_5,
                 Input_14 := "DB47".Static_6,
                 Input_15 := 25,
                 Input_16 := "DB47".Static_7,
                 InOut_0 := %DB47.DBX1.0,
                 Output_0 => "DB47".Static_0,
                 Output_1 => "DB47".Static_1,
                 Output_2 => "DB47".Static_2);
END_REGION
END_FUNCTION

FUNCTION "FalCmpAlta" : Void   // FC49, LAD
{ S7_Optimized_Access := 'FALSE' }
VERSION : 0.1
   VAR_TEMP   // added for the SCL form of the ladder/FBD networks
      _w1 : Bool;
      _s5time1 : S5Time;
   END_VAR
BEGIN

REGION Network 1